REGION Network 2: Sterowanie grzałką w trybie automatycznym i manualnym
   // Gdy uruchomiony jest tryb automatyczny, wartość temperatury w szklarni powinna się mieścić w zakresie temperatury nastawionej +- wartość histerezy. Gdy jest ona za nieska uruchamiana jest grzałka. W trybie manualnym włączana jest ona od razu po naciśnięciu przycisku do niej przypisanego.
   RUNG wire#powerrail
      Contact( #czy_automatyczny )
      I_Contact( #czy_manualny )
      Sub(in1 := "Tryb_auto_parametry".Temperatura, in2 := #Wartosc_histerezy, out => #Histereza_minus)
      { S7_Templates := "SrcType := Real" } GT_Contact(in1 := #Histereza_minus, in2 := "Wejscia_PLC".Temperatura_wewnetrzna)
      wire#w1
      Coil( "Grzałka" )
   END_RUNG
   RUNG wire#powerrail
      Contact( #czy_manualny )
      I_Contact( #czy_automatyczny )
      Contact( "HMI".Przycisk_grzanie_manual )
   END_RUNG wire#w1
   // the same network as SCL:
   #_w1 := #czy_automatyczny AND NOT #czy_manualny;
   IF #_w1 THEN #Histereza_minus := "Tryb_auto_parametry".Temperatura - #Wartosc_histerezy; END_IF;
   "Grzałka" := (#_w1 AND (#Histereza_minus > "Wejscia_PLC".Temperatura_wewnetrzna)) OR (#czy_manualny AND NOT #czy_automatyczny AND "HMI".Przycisk_grzanie_manual);
END_REGION

REGION Network 3: TO DO Alarmy ostrzegające o nieosiąganiu wymaganej temperatury przez długi czas
   "IEC_Timer_0_DB_2".TON(IN := #czy_automatyczny AND NOT #czy_manualny AND ((#Histereza_plus < "Wejscia_PLC".Temperatura_wewnetrzna) OR (#Histereza_minus > "Wejscia_PLC".Temperatura_wewnetrzna)),
                          PT := T#30m);
   "Alarmy".Warning_wysoka_temp_1 := "IEC_Timer_0_DB_2".Q AND (#Histereza_plus > "Tryb_auto_parametry".Temperatura);
   "Alarmy".Warning_niska_temp_1 := "IEC_Timer_0_DB_2".Q AND (#Histereza_minus < "HMI".Temperatura_auto);
END_REGION
END_FUNCTION

FUNCTION "Zapis_parametrow_trybu_auto" : Void   // FC4, LAD
{ S7_Optimized_Access := 'TRUE' }
VERSION : 0.1
BEGIN

REGION Network 1: Zapis wybranych na HMI parametrów, aby zostały one stałe do kolejnego zatwierdzenia ich zmiany.
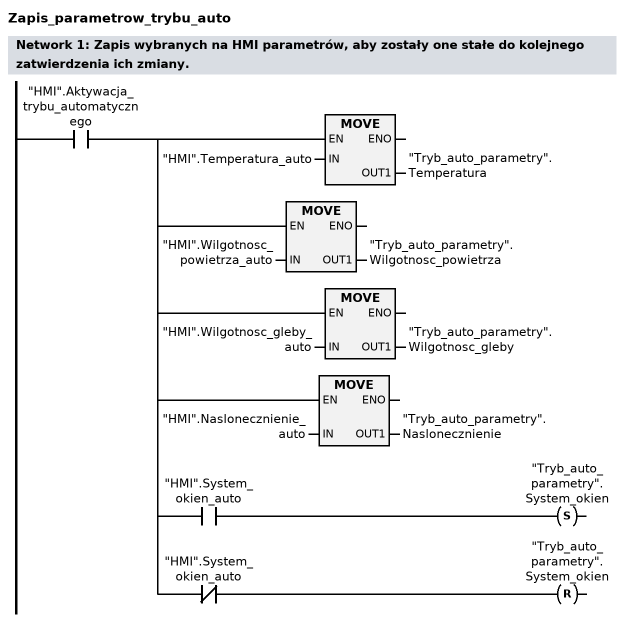
   RUNG wire#powerrail
      Contact( "HMI".Aktywacja_trybu_automatycznego )
      wire#w1
      Move(in := "HMI".Temperatura_auto, out1 => "Tryb_auto_parametry".Temperatura)
   END_RUNG
   RUNG wire#w1
      Move(in := "HMI".Wilgotnosc_powietrza_auto, out1 => "Tryb_auto_parametry".Wilgotnosc_powietrza)
   END_RUNG
   RUNG wire#w1
      Move(in := "HMI".Wilgotnosc_gleby_auto, out1 => "Tryb_auto_parametry".Wilgotnosc_gleby)
   END_RUNG
   RUNG wire#w1
      Move(in := "HMI".Naslonecznienie_auto, out1 => "Tryb_auto_parametry".Naslonecznienie)
   END_RUNG
   RUNG wire#w1
      Contact( "HMI".System_okien_auto )
      S_Coil( "Tryb_auto_parametry".System_okien )
   END_RUNG
   RUNG wire#w1
      I_Contact( "HMI".System_okien_auto )
      R_Coil( "Tryb_auto_parametry".System_okien )
   END_RUNG
   // the same network as SCL:
   IF "HMI".Aktywacja_trybu_automatycznego THEN
       "Tryb_auto_parametry".Temperatura := "HMI".Temperatura_auto;
       "Tryb_auto_parametry".Wilgotnosc_powietrza := "HMI".Wilgotnosc_powietrza_auto;
       "Tryb_auto_parametry".Wilgotnosc_gleby := "HMI".Wilgotnosc_gleby_auto;
       "Tryb_auto_parametry".Naslonecznienie := "HMI".Naslonecznienie_auto;
   END_IF;
   IF "HMI".Aktywacja_trybu_automatycznego AND "HMI".System_okien_auto THEN
       "Tryb_auto_parametry".System_okien := TRUE;
   END_IF;
   IF "HMI".Aktywacja_trybu_automatycznego AND NOT "HMI".System_okien_auto THEN
       "Tryb_auto_parametry".System_okien := FALSE;
   END_IF;
END_REGION
END_FUNCTION

FUNCTION "Jaki_Tryb" : Void   // FC5, LAD
{ S7_Optimized_Access := 'TRUE' }
VERSION : 0.1
BEGIN

REGION Network 1: Reset trybu auto jesli wykryje jakikolwiek inny tryb
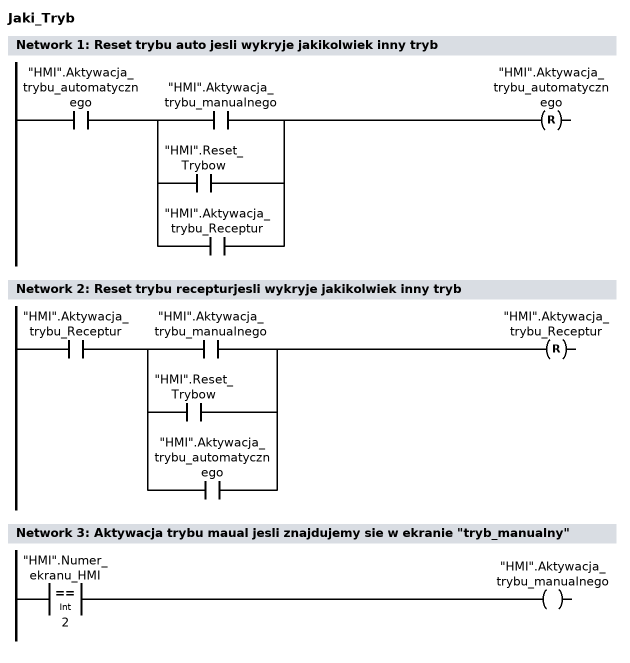
   RUNG wire#powerrail
      Contact( "HMI".Aktywacja_trybu_automatycznego )
      wire#w1
      Contact( "HMI".Aktywacja_trybu_manualnego )
      wire#w2
      R_Coil( "HMI".Aktywacja_trybu_automatycznego )
   END_RUNG
   RUNG wire#w1
      Contact( "HMI".Reset_Trybow )
   END_RUNG wire#w2
   RUNG wire#w1
      Contact( "HMI".Aktywacja_trybu_Receptur )
   END_RUNG wire#w2
   // the same network as SCL:
   IF "HMI".Aktywacja_trybu_automatycznego AND ("HMI".Aktywacja_trybu_manualnego OR "HMI".Reset_Trybow OR "HMI".Aktywacja_trybu_Receptur) THEN
       "HMI".Aktywacja_trybu_automatycznego := FALSE;
   END_IF;
END_REGION

REGION Network 2: Reset trybu recepturjesli wykryje jakikolwiek inny tryb
   RUNG wire#powerrail
      Contact( "HMI".Aktywacja_trybu_Receptur )
      wire#w1
      Contact( "HMI".Aktywacja_trybu_manualnego )
      wire#w2
      R_Coil( "HMI".Aktywacja_trybu_Receptur )
   END_RUNG
   RUNG wire#w1
      Contact( "HMI".Reset_Trybow )
   END_RUNG wire#w2
   RUNG wire#w1
      Contact( "HMI".Aktywacja_trybu_automatycznego )
   END_RUNG wire#w2
   // the same network as SCL:
   IF "HMI".Aktywacja_trybu_Receptur AND ("HMI".Aktywacja_trybu_manualnego OR "HMI".Reset_Trybow OR "HMI".Aktywacja_trybu_automatycznego) THEN
       "HMI".Aktywacja_trybu_Receptur := FALSE;
   END_IF;
END_REGION

REGION Network 3: Aktywacja trybu maual jesli znajdujemy sie w ekranie "tryb_manualny"
   RUNG wire#powerrail
      { S7_Templates := "SrcType := Int" } EQ_Contact(in1 := "HMI".Numer_ekranu_HMI, in2 := 2)
      Coil( "HMI".Aktywacja_trybu_manualnego )
   END_RUNG
   // the same network as SCL:
   "HMI".Aktywacja_trybu_manualnego := "HMI".Numer_ekranu_HMI = 2;
END_REGION
END_FUNCTION

FUNCTION "Ograniczanie_wartosci_parametrow" : Void   // FC6, LAD
TITLE = Każdy z poniższych network-ów odpowiada za to, aby po ustawieniu na HMI wartości przekraczajacej dopuszczalną, ta pozostała w wymaganym zakresie.
{ S7_Optimized_Access := 'TRUE' }
VERSION : 0.1
BEGIN

REGION Network 1: Ograniczenie dla wartosci ustawionej temperatury w trybie automatycznym
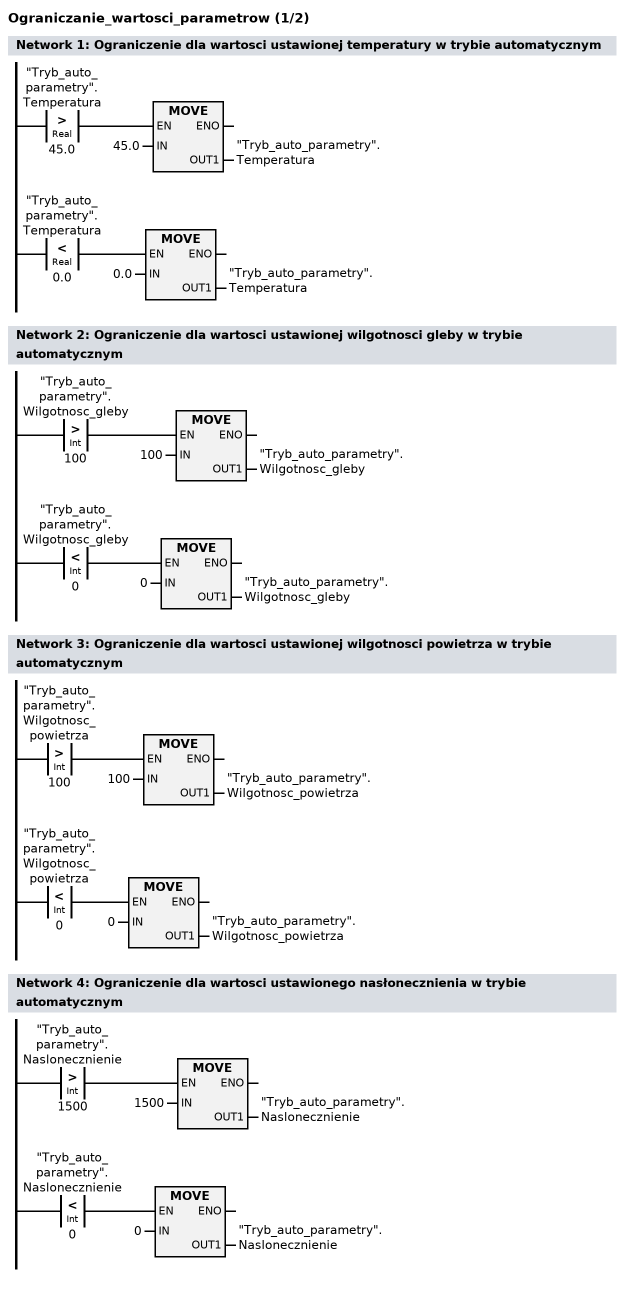
   RUNG wire#powerrail
      { S7_Templates := "SrcType := Real" } GT_Contact(in1 := "Tryb_auto_parametry".Temperatura, in2 := 45.0)
      Move(in := 45.0, out1 => "Tryb_auto_parametry".Temperatura)
   END_RUNG
   RUNG wire#powerrail
      { S7_Templates := "SrcType := Real" } LT_Contact(in1 := "Tryb_auto_parametry".Temperatura, in2 := 0.0)
      Move(in := 0.0, out1 => "Tryb_auto_parametry".Temperatura)
   END_RUNG
   // the same network as SCL:
   IF "Tryb_auto_parametry".Temperatura > 45.0 THEN "Tryb_auto_parametry".Temperatura := 45.0; END_IF;
   IF "Tryb_auto_parametry".Temperatura < 0.0 THEN "Tryb_auto_parametry".Temperatura := 0.0; END_IF;
END_REGION

REGION Network 2: Ograniczenie dla wartosci ustawionej wilgotnosci gleby w trybie automatycznym
   RUNG wire#powerrail
      { S7_Templates := "SrcType := Int" } GT_Contact(in1 := "Tryb_auto_parametry".Wilgotnosc_gleby, in2 := 100)
      Move(in := 100, out1 => "Tryb_auto_parametry".Wilgotnosc_gleby)
   END_RUNG
   RUNG wire#powerrail
      { S7_Templates := "SrcType := Int" } LT_Contact(in1 := "Tryb_auto_parametry".Wilgotnosc_gleby, in2 := 0)
      Move(in := 0, out1 => "Tryb_auto_parametry".Wilgotnosc_gleby)
   END_RUNG
   // the same network as SCL:
   IF "Tryb_auto_parametry".Wilgotnosc_gleby > 100 THEN
       "Tryb_auto_parametry".Wilgotnosc_gleby := 100;
   END_IF;
   IF "Tryb_auto_parametry".Wilgotnosc_gleby < 0 THEN "Tryb_auto_parametry".Wilgotnosc_gleby := 0; END_IF;
END_REGION

REGION Network 3: Ograniczenie dla wartosci ustawionej wilgotnosci powietrza w trybie automatycznym
   RUNG wire#powerrail
      { S7_Templates := "SrcType := Int" } GT_Contact(in1 := "Tryb_auto_parametry".Wilgotnosc_powietrza, in2 := 100)
      Move(in := 100, out1 => "Tryb_auto_parametry".Wilgotnosc_powietrza)
   END_RUNG
   RUNG wire#powerrail
      { S7_Templates := "SrcType := Int" } LT_Contact(in1 := "Tryb_auto_parametry".Wilgotnosc_powietrza, in2 := 0)
      Move(in := 0, out1 => "Tryb_auto_parametry".Wilgotnosc_powietrza)
   END_RUNG
   // the same network as SCL:
   IF "Tryb_auto_parametry".Wilgotnosc_powietrza > 100 THEN
       "Tryb_auto_parametry".Wilgotnosc_powietrza := 100;
   END_IF;
   IF "Tryb_auto_parametry".Wilgotnosc_powietrza < 0 THEN
       "Tryb_auto_parametry".Wilgotnosc_powietrza := 0;
   END_IF;
END_REGION

REGION Network 4: Ograniczenie dla wartosci ustawionego nasłonecznienia w trybie automatycznym
   RUNG wire#powerrail
      { S7_Templates := "SrcType := Int" } GT_Contact(in1 := "Tryb_auto_parametry".Naslonecznienie, in2 := 1500)
      Move(in := 1500, out1 => "Tryb_auto_parametry".Naslonecznienie)
   END_RUNG
   RUNG wire#powerrail
      { S7_Templates := "SrcType := Int" } LT_Contact(in1 := "Tryb_auto_parametry".Naslonecznienie, in2 := 0)
      Move(in := 0, out1 => "Tryb_auto_parametry".Naslonecznienie)
   END_RUNG
   // the same network as SCL:
   IF "Tryb_auto_parametry".Naslonecznienie > 1500 THEN
       "Tryb_auto_parametry".Naslonecznienie := 1500;
   END_IF;
   IF "Tryb_auto_parametry".Naslonecznienie < 0 THEN "Tryb_auto_parametry".Naslonecznienie := 0; END_IF;
END_REGION

REGION Network 5: Ograniczenie dla wartosci ustawionego stężenia CO2 w trybie automatycznym
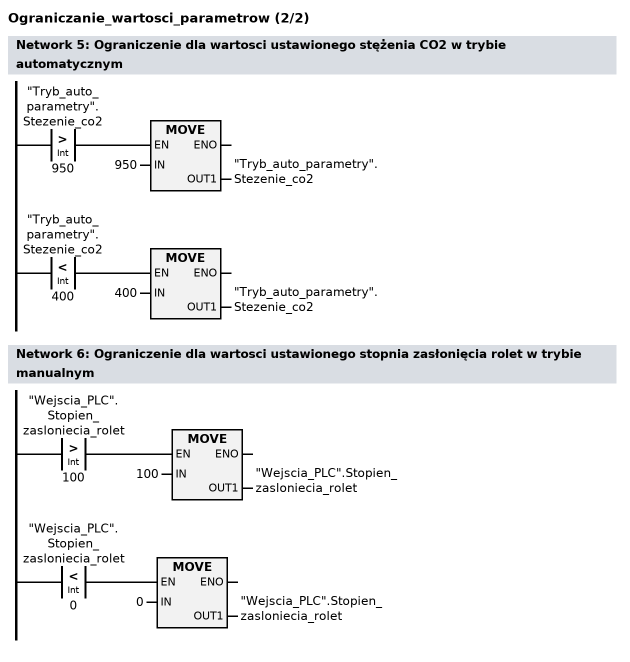
   RUNG wire#powerrail
      { S7_Templates := "SrcType := Int" } GT_Contact(in1 := "Tryb_auto_parametry".Stezenie_co2, in2 := 950)
      Move(in := 950, out1 => "Tryb_auto_parametry".Stezenie_co2)
   END_RUNG
   RUNG wire#powerrail
      { S7_Templates := "SrcType := Int" } LT_Contact(in1 := "Tryb_auto_parametry".Stezenie_co2, in2 := 400)
      Move(in := 400, out1 => "Tryb_auto_parametry".Stezenie_co2)
   END_RUNG
   // the same network as SCL:
   IF "Tryb_auto_parametry".Stezenie_co2 > 950 THEN "Tryb_auto_parametry".Stezenie_co2 := 950; END_IF;
   IF "Tryb_auto_parametry".Stezenie_co2 < 400 THEN "Tryb_auto_parametry".Stezenie_co2 := 400; END_IF;
END_REGION

REGION Network 6: Ograniczenie dla wartosci ustawionego stopnia zasłonięcia rolet w trybie manualnym
   RUNG wire#powerrail
      { S7_Templates := "SrcType := Int" } GT_Contact(in1 := "Wejscia_PLC".Stopien_zasloniecia_rolet, in2 := 100)
      Move(in := 100, out1 => "Wejscia_PLC".Stopien_zasloniecia_rolet)
   END_RUNG
   RUNG wire#powerrail
      { S7_Templates := "SrcType := Int" } LT_Contact(in1 := "Wejscia_PLC".Stopien_zasloniecia_rolet, in2 := 0)
      Move(in := 0, out1 => "Wejscia_PLC".Stopien_zasloniecia_rolet)
   END_RUNG
   // the same network as SCL:
   IF "Wejscia_PLC".Stopien_zasloniecia_rolet > 100 THEN
       "Wejscia_PLC".Stopien_zasloniecia_rolet := 100;
   END_IF;
   IF "Wejscia_PLC".Stopien_zasloniecia_rolet < 0 THEN "Wejscia_PLC".Stopien_zasloniecia_rolet := 0; END_IF;
END_REGION
END_FUNCTION

FUNCTION "Sterowanie_podlewaniem_zraszaniem" : Void   // FC7, LAD
{ S7_Optimized_Access := 'TRUE' }
VERSION : 0.1
   VAR_INPUT
      Czy_automatyczny : Bool;
      Czy_manualny : Bool;
   END_VAR
BEGIN

REGION Network 1: Sterowanie pompą zraszaczy, które odpowiadają za wilgotność powietrza w szklarni
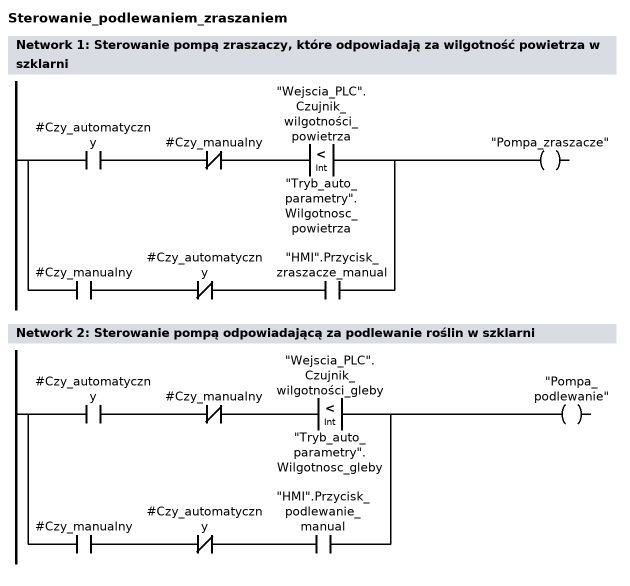
   RUNG wire#powerrail
      Contact( #Czy_automatyczny )
      I_Contact( #Czy_manualny )
      { S7_Templates := "SrcType := Int" } LT_Contact(in1 := "Wejscia_PLC".Czujnik_wilgotności_powietrza, in2 := "Tryb_auto_parametry".Wilgotnosc_powietrza)
      wire#w1
      Coil( "Pompa_zraszacze" )
   END_RUNG
   RUNG wire#powerrail
      Contact( #Czy_manualny )
      I_Contact( #Czy_automatyczny )
      Contact( "HMI".Przycisk_zraszacze_manual )
   END_RUNG wire#w1
   // the same network as SCL:
   "Pompa_zraszacze" := (#Czy_automatyczny AND NOT #Czy_manualny AND ("Wejscia_PLC".Czujnik_wilgotności_powietrza < "Tryb_auto_parametry".Wilgotnosc_powietrza)) OR (#Czy_manualny AND NOT #Czy_automatyczny AND "HMI".Przycisk_zraszacze_manual);
END_REGION

REGION Network 2: Sterowanie pompą odpowiadającą za podlewanie roślin w szklarni
   RUNG wire#powerrail
      Contact( #Czy_automatyczny )
      I_Contact( #Czy_manualny )
      { S7_Templates := "SrcType := Int" } LT_Contact(in1 := "Wejscia_PLC".Czujnik_wilgotności_gleby, in2 := "Tryb_auto_parametry".Wilgotnosc_gleby)
      wire#w1
      Coil( "Pompa_podlewanie" )
   END_RUNG
   RUNG wire#powerrail
      Contact( #Czy_manualny )
      I_Contact( #Czy_automatyczny )
      Contact( "HMI".Przycisk_podlewanie_manual )
   END_RUNG wire#w1
   // the same network as SCL:
   "Pompa_podlewanie" := (#Czy_automatyczny AND NOT #Czy_manualny AND ("Wejscia_PLC".Czujnik_wilgotności_gleby < "Tryb_auto_parametry".Wilgotnosc_gleby)) OR (#Czy_manualny AND NOT #Czy_automatyczny AND "HMI".Przycisk_podlewanie_manual);
END_REGION
END_FUNCTION

FUNCTION "Sterowanie_oknami" : Void   // FC8, LAD
{ S7_Optimized_Access := 'TRUE' }
VERSION : 0.1
   VAR_INPUT
      czy_manualny : Bool;
      czy_automatyczny : Bool;
   END_VAR
   VAR_TEMP
      Histereza_plus : Int;
      Histereza_minus : Int;
      Zakres_temp_gora : Real;   // Górny zakres temperatury zewnętrznej dla której w trybie automatycznym będą otwierane okna
      Zakres_temp_dol : Real;   // Dolny zakres temperatury zewnętrznej dla której w trybie automatycznym będą otwierane okna
   END_VAR
   VAR CONSTANT
      Histereza : Int := 25;   // Histereza, która określa kiedy stan CO2 w szklarni jest uznawany za prawidłowy
   END_VAR
BEGIN

REGION Network 1: Operacje matematyczne używane w networku 2. i 3.
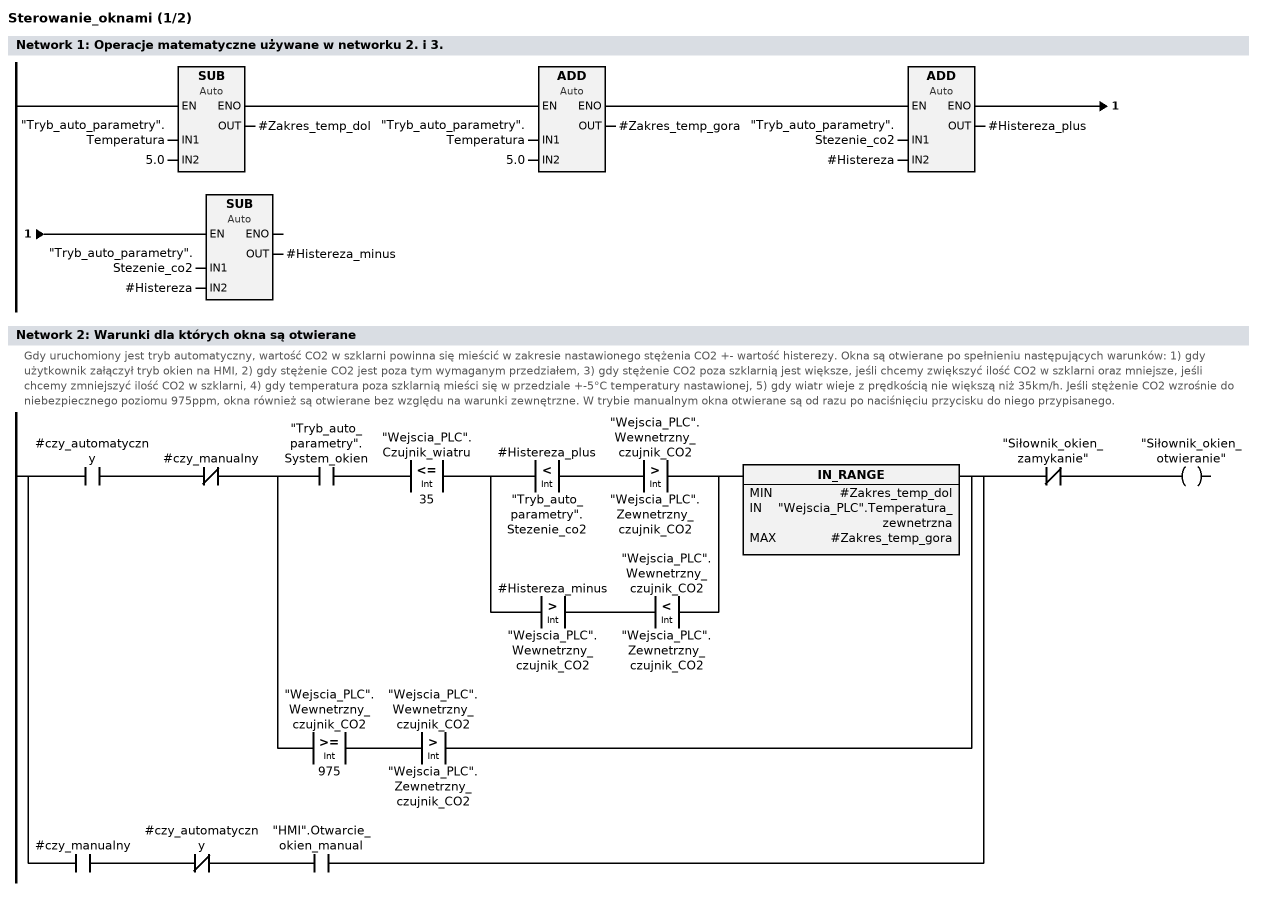
   RUNG wire#powerrail
      Sub(in1 := "Tryb_auto_parametry".Temperatura, in2 := 5.0, out => #Zakres_temp_dol)
      Add(in1 := "Tryb_auto_parametry".Temperatura, in2 := 5.0, out => #Zakres_temp_gora)
      Add(in1 := "Tryb_auto_parametry".Stezenie_co2, in2 := #Histereza, out => #Histereza_plus)
      Sub(in1 := "Tryb_auto_parametry".Stezenie_co2, in2 := #Histereza, out => #Histereza_minus)
   END_RUNG
   // the same network as SCL:
   #Zakres_temp_dol := "Tryb_auto_parametry".Temperatura - 5.0;
   #Zakres_temp_gora := "Tryb_auto_parametry".Temperatura + 5.0;
   #Histereza_plus := "Tryb_auto_parametry".Stezenie_co2 + #Histereza;
   #Histereza_minus := "Tryb_auto_parametry".Stezenie_co2 - #Histereza;
END_REGION

REGION Network 2: Warunki dla których okna są otwierane
   // Gdy uruchomiony jest tryb automatyczny, wartość CO2 w szklarni powinna się mieścić w zakresie nastawionego stężenia CO2 +- wartość histerezy. Okna są otwierane po spełnieniu następujących warunków: 1) gdy użytkownik załączył tryb okien na HMI, 2) gdy stężenie CO2 jest poza tym wymaganym przedziałem, 3) gdy stężenie CO2 poza szklarnią jest większe, jeśli chcemy zwiększyć ilość CO2 w szklarni oraz mniejsze, jeśli chcemy zmniejszyć ilość CO2 w szklarni, 4) gdy temperatura poza szklarnią mieści się w przedziale +-5°C temperatury nastawionej, 5) gdy wiatr wieje z prędkością nie większą niż 35km/h. Jeśli stężenie CO2 wzrośnie do niebezpiecznego poziomu 975ppm, okna również są otwierane bez względu na warunki zewnętrzne. W trybie manualnym okna otwierane są od razu po naciśnięciu przycisku do niego przypisanego.
   RUNG wire#powerrail
      Contact( #czy_automatyczny )
      I_Contact( #czy_manualny )
      wire#w1
      Contact( "Tryb_auto_parametry".System_okien )
      { S7_Templates := "SrcType := Int" } LE_Contact(in1 := "Wejscia_PLC".Czujnik_wiatru, in2 := 35)
      wire#w2
      { S7_Templates := "SrcType := Int" } LT_Contact(in1 := #Histereza_plus, in2 := "Tryb_auto_parametry".Stezenie_co2)
      { S7_Templates := "SrcType := Int" } GT_Contact(in1 := "Wejscia_PLC".Wewnetrzny_czujnik_CO2, in2 := "Wejscia_PLC".Zewnetrzny_czujnik_CO2)
      wire#w3
      { S7_Templates := "SrcType := Real" } InRange(min := #Zakres_temp_dol, in := "Wejscia_PLC".Temperatura_zewnetrzna, max := #Zakres_temp_gora)
      wire#w4
      I_Contact( "Siłownik_okien_zamykanie" )
      Coil( "Siłownik_okien_otwieranie" )
   END_RUNG
   RUNG wire#w2
      { S7_Templates := "SrcType := Int" } GT_Contact(in1 := #Histereza_minus, in2 := "Wejscia_PLC".Wewnetrzny_czujnik_CO2)
      { S7_Templates := "SrcType := Int" } LT_Contact(in1 := "Wejscia_PLC".Wewnetrzny_czujnik_CO2, in2 := "Wejscia_PLC".Zewnetrzny_czujnik_CO2)
   END_RUNG wire#w3
   RUNG wire#w1
      { S7_Templates := "SrcType := Int" } GE_Contact(in1 := "Wejscia_PLC".Wewnetrzny_czujnik_CO2, in2 := 975)
      { S7_Templates := "SrcType := Int" } GT_Contact(in1 := "Wejscia_PLC".Wewnetrzny_czujnik_CO2, in2 := "Wejscia_PLC".Zewnetrzny_czujnik_CO2)
   END_RUNG wire#w4
   RUNG wire#powerrail
      Contact( #czy_manualny )
      I_Contact( #czy_automatyczny )
      Contact( "HMI".Otwarcie_okien_manual )
   END_RUNG wire#w4
   // the same network as SCL:
   "Siłownik_okien_otwieranie" := ((#czy_automatyczny AND NOT #czy_manualny AND (("Tryb_auto_parametry".System_okien AND ("Wejscia_PLC".Czujnik_wiatru <= 35) AND (((#Histereza_plus < "Tryb_auto_parametry".Stezenie_co2) AND ("Wejscia_PLC".Wewnetrzny_czujnik_CO2 > "Wejscia_PLC".Zewnetrzny_czujnik_CO2)) OR ((#Histereza_minus > "Wejscia_PLC".Wewnetrzny_czujnik_CO2) AND ("Wejscia_PLC".Wewnetrzny_czujnik_CO2 < "Wejscia_PLC".Zewnetrzny_czujnik_CO2))) AND (#Zakres_temp_dol <= "Wejscia_PLC".Temperatura_zewnetrzna) AND ("Wejscia_PLC".Temperatura_zewnetrzna <= #Zakres_temp_gora)) OR (("Wejscia_PLC".Wewnetrzny_czujnik_CO2 >= 975) AND ("Wejscia_PLC".Wewnetrzny_czujnik_CO2 > "Wejscia_PLC".Zewnetrzny_czujnik_CO2)))) OR (#czy_manualny AND NOT #czy_automatyczny AND "HMI".Otwarcie_okien_manual)) AND NOT "Siłownik_okien_zamykanie";
END_REGION

REGION Network 3: Warunki dla których okna są zamykane
   // W trybie automatycznym okna są zamykane: 1) gdy tryb okien został wyłączony przez użytkownika, 2) gdy stężenie CO2 w szklarni wynosi zadaną wartość tego parametru +- histereza, 3) gdy stężenie CO2 poza szklarnią jest mniejsze, niż wewnątrz, jeśli chcemy zwiększyć jego ilość oraz większe, gdy chcemy zmniejszyć jego ilość, 4) gdy tempperatura zewnętrzna różni się o ponad 5°C od zadanej, 5) gdy wiatr wieje z prędkością większą niż 35km/h, 6) gdy stężenie CO2 w szklarni nie przekracza 955ppm lub przekracza, ale stężenie CO2 poza szklarnią jest większe. W trybie manualnym okna są zamykane, gdy przełączk na HMI znajdzie się w pozycji "ZAMKNIĘTE".
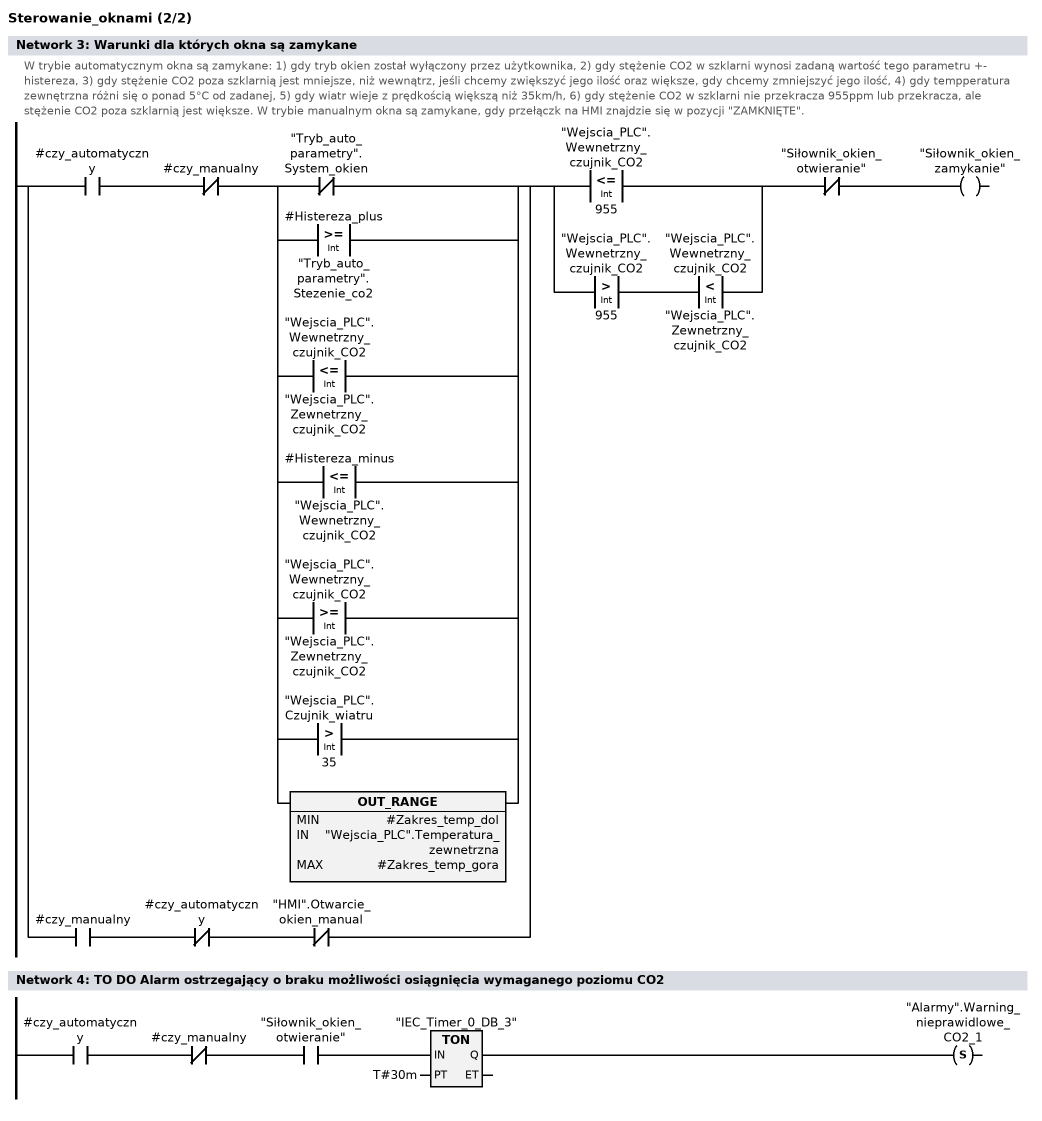
   "Siłownik_okien_zamykanie" := ((#czy_automatyczny AND NOT #czy_manualny AND (NOT "Tryb_auto_parametry".System_okien OR (#Histereza_plus >= "Tryb_auto_parametry".Stezenie_co2) OR ("Wejscia_PLC".Wewnetrzny_czujnik_CO2 <= "Wejscia_PLC".Zewnetrzny_czujnik_CO2) OR (#Histereza_minus <= "Wejscia_PLC".Wewnetrzny_czujnik_CO2) OR ("Wejscia_PLC".Wewnetrzny_czujnik_CO2 >= "Wejscia_PLC".Zewnetrzny_czujnik_CO2) OR ("Wejscia_PLC".Czujnik_wiatru > 35) OR ("Wejscia_PLC".Temperatura_zewnetrzna < #Zakres_temp_dol) OR ("Wejscia_PLC".Temperatura_zewnetrzna > #Zakres_temp_gora))) OR (#czy_manualny AND NOT #czy_automatyczny AND NOT "HMI".Otwarcie_okien_manual)) AND (("Wejscia_PLC".Wewnetrzny_czujnik_CO2 <= 955) OR (("Wejscia_PLC".Wewnetrzny_czujnik_CO2 > 955) AND ("Wejscia_PLC".Wewnetrzny_czujnik_CO2 < "Wejscia_PLC".Zewnetrzny_czujnik_CO2))) AND NOT "Siłownik_okien_otwieranie";
END_REGION

REGION Network 4: TO DO Alarm ostrzegający o braku możliwości osiągnięcia wymaganego poziomu CO2
   "IEC_Timer_0_DB_3".TON(IN := #czy_automatyczny AND NOT #czy_manualny AND "Siłownik_okien_otwieranie",
                          PT := T#30m);
   IF "IEC_Timer_0_DB_3".Q THEN "Alarmy".Warning_nieprawidlowe_CO2_1 := TRUE; END_IF;
END_REGION
END_FUNCTION

FUNCTION "SYMULACJA" : Void   // FC9, LAD
{ S7_Optimized_Access := 'TRUE' }
VERSION : 0.1
   VAR_INPUT
      counters : Bool;
   END_VAR
   VAR_TEMP
      temperatura_temp : Real;
      roznica_temperatur : Real;
      "wilgotność powietrza_temp" : Int;
      wilgotnosc_gleby_temp : Int;
      stezenie_CO2 : Int;
      natezenie_swiatla_temp : Int;
      odsloniecie_okna_temp : Real;
      pedkosc_wiatru_temp : Real;
      rand : Real;
      error : Bool;
      status : Int;
      sub_status : Int;
      rolety_temp : Real;
      test1 : Real;
   END_VAR
   VAR_TEMP   // added for the SCL form of the ladder/FBD networks
      _w1 : Bool;
   END_VAR
BEGIN

REGION Network 1: blok oblicza roznice temperatur
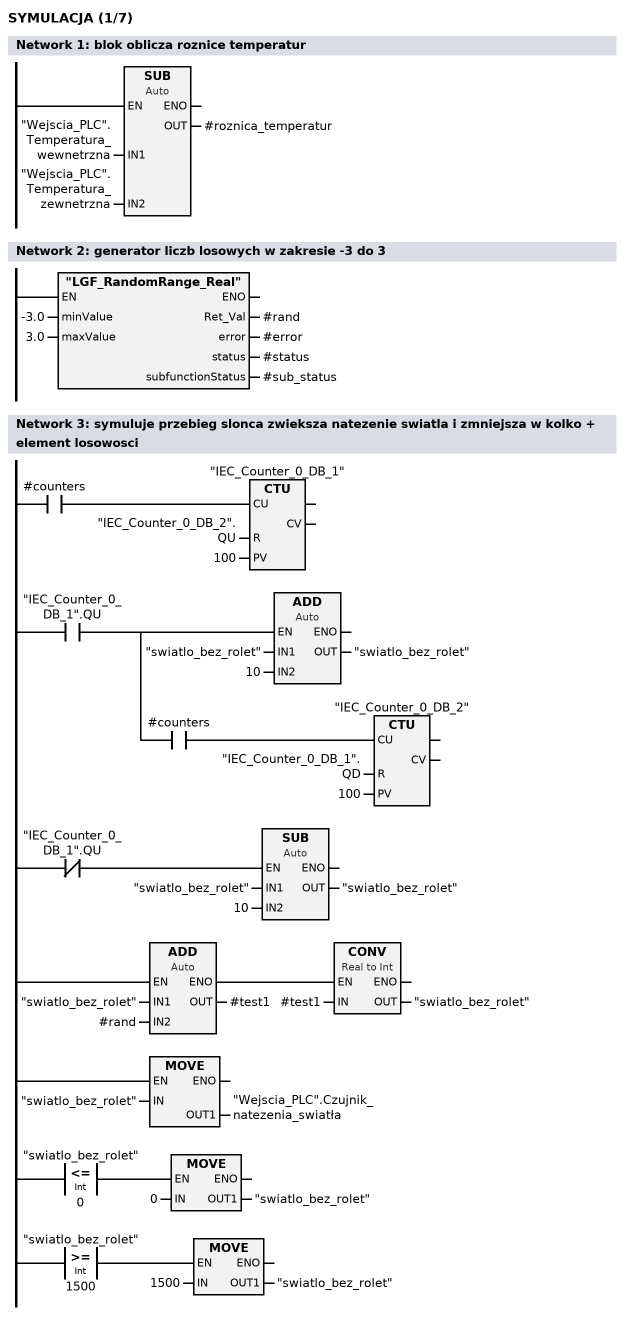
   RUNG wire#powerrail
      { S7_GenerateENO := "TRUE" } Sub(in1 := "Wejscia_PLC".Temperatura_wewnetrzna, in2 := "Wejscia_PLC".Temperatura_zewnetrzna, out => #roznica_temperatur)
   END_RUNG
   // the same network as SCL:
   #roznica_temperatur := "Wejscia_PLC".Temperatura_wewnetrzna - "Wejscia_PLC".Temperatura_zewnetrzna;
END_REGION

REGION Network 2: generator liczb losowych w zakresie -3 do 3
   RUNG wire#powerrail
      "LGF_RandomRange_Real"(minValue := -3.0, maxValue := 3.0, Ret_Val => #rand, error => #error, status => #status, subfunctionStatus => #sub_status)
   END_RUNG
   // the same network as SCL:
   #rand := "LGF_RandomRange_Real"(minValue := -3.0,
                           maxValue := 3.0,
                           error => #error,
                           status => #status,
                           subfunctionStatus => #sub_status);
END_REGION

REGION Network 3: symuluje przebieg slonca zwieksza natezenie swiatla i zmniejsza w kolko + element losowosci
   // ENO of a box is taken as its EN; it also drops when the box reports an error
   "IEC_Counter_0_DB_1".CTU(CU := #counters, R := "IEC_Counter_0_DB_2".QU, PV := 100);
   IF "IEC_Counter_0_DB_1".QU THEN "swiatlo_bez_rolet" := "swiatlo_bez_rolet" + 10; END_IF;
   "IEC_Counter_0_DB_2".CTU(CU := "IEC_Counter_0_DB_1".QU AND #counters,
                           R := "IEC_Counter_0_DB_1".QD,
                           PV := 100);
   IF NOT "IEC_Counter_0_DB_1".QU THEN "swiatlo_bez_rolet" := "swiatlo_bez_rolet" - 10; END_IF;
   #test1 := "swiatlo_bez_rolet" + #rand;
   "swiatlo_bez_rolet" := REAL_TO_INT(#test1);
   "Wejscia_PLC".Czujnik_natezenia_swiatła := "swiatlo_bez_rolet";
   IF "swiatlo_bez_rolet" <= 0 THEN "swiatlo_bez_rolet" := 0; END_IF;
   IF "swiatlo_bez_rolet" >= 1500 THEN "swiatlo_bez_rolet" := 1500; END_IF;
END_REGION

REGION Network 4: funkcja oblicza liniową zależność natężenia światła od zasłonięcia rolet
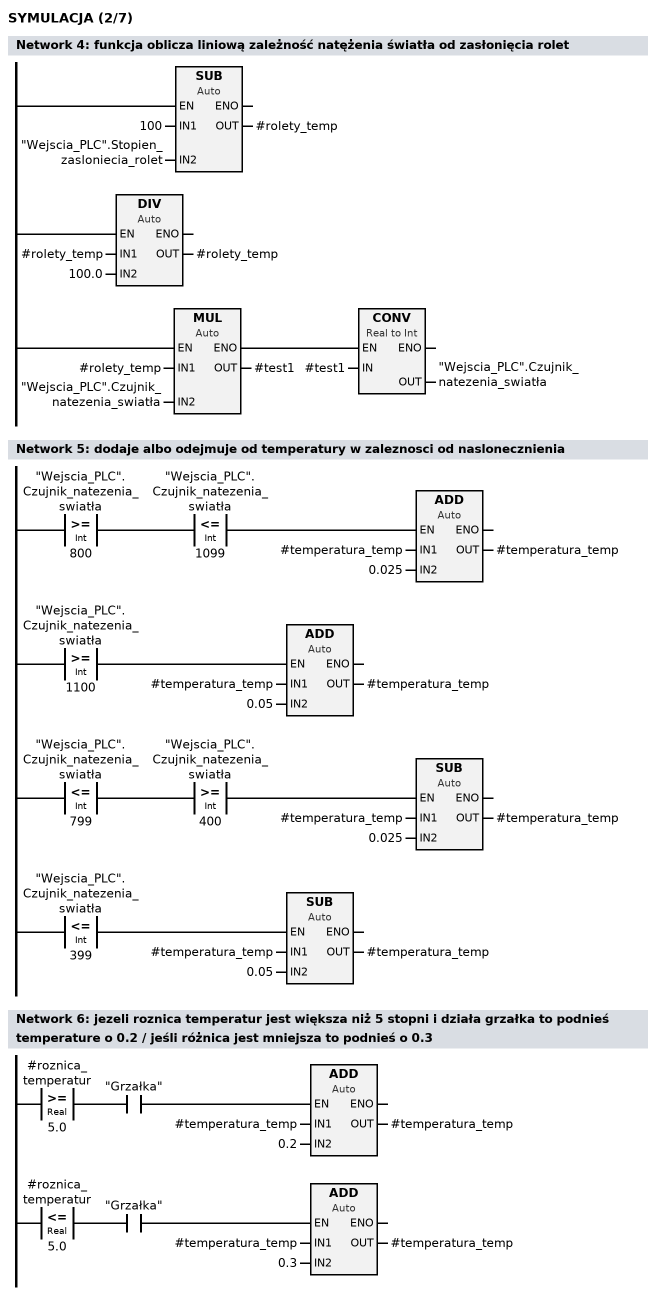
   RUNG wire#powerrail
      { S7_GenerateENO := "TRUE" } Sub(in1 := 100, in2 := "Wejscia_PLC".Stopien_zasloniecia_rolet, out => #rolety_temp)
   END_RUNG
   RUNG wire#powerrail
      { S7_GenerateENO := "TRUE" } Div(in1 := #rolety_temp, in2 := 100.0, out => #rolety_temp)
   END_RUNG
   RUNG wire#powerrail
      { S7_GenerateENO := "TRUE" } Mul(in1 := #rolety_temp, in2 := "Wejscia_PLC".Czujnik_natezenia_swiatła, out => #test1)
      { S7_Templates := "[SrcType := Real, DestType := Int]"; S7_GenerateENO := "TRUE" } Convert(in := #test1, out => "Wejscia_PLC".Czujnik_natezenia_swiatła)
   END_RUNG
   // the same network as SCL:
   // ENO of a box is taken as its EN; it also drops when the box reports an error
   #rolety_temp := 100 - "Wejscia_PLC".Stopien_zasloniecia_rolet;
   #rolety_temp := #rolety_temp / 100.0;
   #test1 := #rolety_temp * "Wejscia_PLC".Czujnik_natezenia_swiatła;
   "Wejscia_PLC".Czujnik_natezenia_swiatła := REAL_TO_INT(#test1);
END_REGION

REGION Network 5: dodaje albo odejmuje od temperatury w zaleznosci od naslonecznienia
   RUNG wire#powerrail
      { S7_Templates := "SrcType := Int" } GE_Contact(in1 := "Wejscia_PLC".Czujnik_natezenia_swiatła, in2 := 800)
      { S7_Templates := "SrcType := Int" } LE_Contact(in1 := "Wejscia_PLC".Czujnik_natezenia_swiatła, in2 := 1099)
      { S7_GenerateENO := "TRUE" } Add(in1 := #temperatura_temp, in2 := 0.025, out => #temperatura_temp)
   END_RUNG
   RUNG wire#powerrail
      { S7_Templates := "SrcType := Int" } GE_Contact(in1 := "Wejscia_PLC".Czujnik_natezenia_swiatła, in2 := 1100)
      { S7_GenerateENO := "TRUE" } Add(in1 := #temperatura_temp, in2 := 0.05, out => #temperatura_temp)
   END_RUNG
   RUNG wire#powerrail
      { S7_Templates := "SrcType := Int" } LE_Contact(in1 := "Wejscia_PLC".Czujnik_natezenia_swiatła, in2 := 799)
      { S7_Templates := "SrcType := Int" } GE_Contact(in1 := "Wejscia_PLC".Czujnik_natezenia_swiatła, in2 := 400)
      { S7_GenerateENO := "TRUE" } Sub(in1 := #temperatura_temp, in2 := 0.025, out => #temperatura_temp)
   END_RUNG
   RUNG wire#powerrail
      { S7_Templates := "SrcType := Int" } LE_Contact(in1 := "Wejscia_PLC".Czujnik_natezenia_swiatła, in2 := 399)
      { S7_GenerateENO := "TRUE" } Sub(in1 := #temperatura_temp, in2 := 0.05, out => #temperatura_temp)
   END_RUNG
   // the same network as SCL:
   IF ("Wejscia_PLC".Czujnik_natezenia_swiatła >= 800) AND ("Wejscia_PLC".Czujnik_natezenia_swiatła <= 1099) THEN
       #temperatura_temp := #temperatura_temp + 0.025;
   END_IF;
   IF "Wejscia_PLC".Czujnik_natezenia_swiatła >= 1100 THEN
       #temperatura_temp := #temperatura_temp + 0.05;
   END_IF;
   IF ("Wejscia_PLC".Czujnik_natezenia_swiatła <= 799) AND ("Wejscia_PLC".Czujnik_natezenia_swiatła >= 400) THEN
       #temperatura_temp := #temperatura_temp - 0.025;
   END_IF;
   IF "Wejscia_PLC".Czujnik_natezenia_swiatła <= 399 THEN
       #temperatura_temp := #temperatura_temp - 0.05;
   END_IF;
END_REGION

REGION Network 6: jezeli roznica temperatur jest większa niż 5 stopni i działa grzałka to podnieś temperature o 0.2 / jeśli różnica jest mniejsza to podnieś o 0.3
   RUNG wire#powerrail
      { S7_Templates := "SrcType := Real" } GE_Contact(in1 := #roznica_temperatur, in2 := 5.0)
      Contact( "Grzałka" )
      { S7_GenerateENO := "TRUE" } Add(in1 := #temperatura_temp, in2 := 0.2, out => #temperatura_temp)
   END_RUNG
   RUNG wire#powerrail
      { S7_Templates := "SrcType := Real" } LE_Contact(in1 := #roznica_temperatur, in2 := 5.0)
      Contact( "Grzałka" )
      { S7_GenerateENO := "TRUE" } Add(in1 := #temperatura_temp, in2 := 0.3, out => #temperatura_temp)
   END_RUNG
   // the same network as SCL:
   IF (#roznica_temperatur >= 5.0) AND "Grzałka" THEN #temperatura_temp := #temperatura_temp + 0.2; END_IF;
   IF (#roznica_temperatur <= 5.0) AND "Grzałka" THEN #temperatura_temp := #temperatura_temp + 0.3; END_IF;
END_REGION

REGION Network 7: jezeli działa wentylator to obniż temperature o 0.1
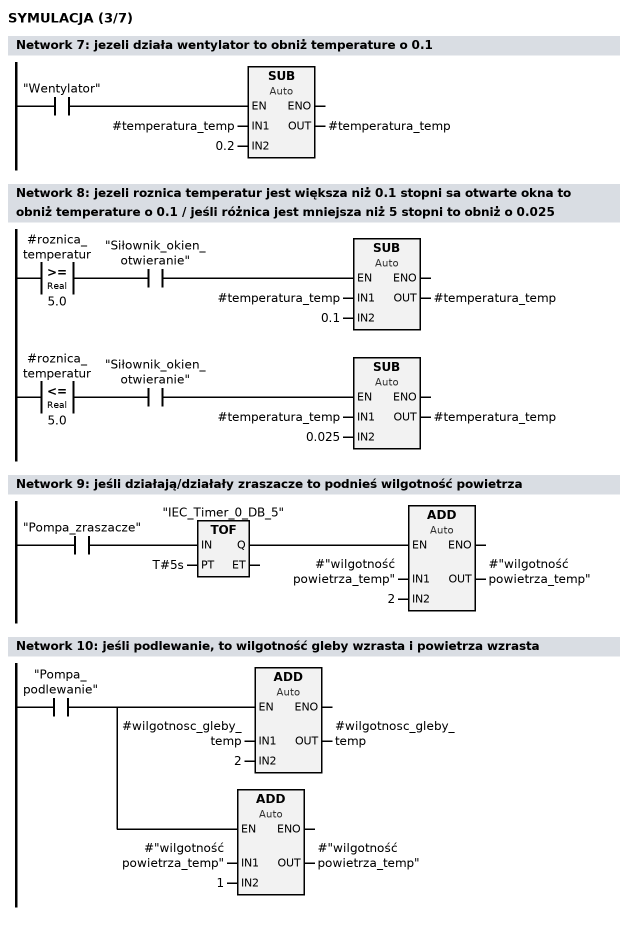
   RUNG wire#powerrail
      Contact( "Wentylator" )
      { S7_GenerateENO := "TRUE" } Sub(in1 := #temperatura_temp, in2 := 0.2, out => #temperatura_temp)
   END_RUNG
   // the same network as SCL:
   IF "Wentylator" THEN #temperatura_temp := #temperatura_temp - 0.2; END_IF;
END_REGION

REGION Network 8: jezeli roznica temperatur jest większa niż 0.1 stopni sa otwarte okna to obniż temperature o 0.1 / jeśli różnica jest mniejsza niż 5 stopni to obniż o 0.025
   RUNG wire#powerrail
      { S7_Templates := "SrcType := Real" } GE_Contact(in1 := #roznica_temperatur, in2 := 5.0)
      Contact( "Siłownik_okien_otwieranie" )
      { S7_GenerateENO := "TRUE" } Sub(in1 := #temperatura_temp, in2 := 0.1, out => #temperatura_temp)
   END_RUNG
   RUNG wire#powerrail
      { S7_Templates := "SrcType := Real" } LE_Contact(in1 := #roznica_temperatur, in2 := 5.0)
      Contact( "Siłownik_okien_otwieranie" )
      { S7_GenerateENO := "TRUE" } Sub(in1 := #temperatura_temp, in2 := 0.025, out => #temperatura_temp)
   END_RUNG
   // the same network as SCL:
   IF (#roznica_temperatur >= 5.0) AND "Siłownik_okien_otwieranie" THEN
       #temperatura_temp := #temperatura_temp - 0.1;
   END_IF;
   IF (#roznica_temperatur <= 5.0) AND "Siłownik_okien_otwieranie" THEN
       #temperatura_temp := #temperatura_temp - 0.025;
   END_IF;
END_REGION

REGION Network 9: jeśli działają/działały zraszacze to podnieś wilgotność powietrza
   "IEC_Timer_0_DB_5".TOF(IN := "Pompa_zraszacze", PT := T#5s);
   IF "IEC_Timer_0_DB_5".Q THEN #"wilgotność powietrza_temp" := #"wilgotność powietrza_temp" + 2; END_IF;
END_REGION

REGION Network 10: jeśli podlewanie, to wilgotność gleby wzrasta i powietrza wzrasta
   RUNG wire#powerrail
      Contact( "Pompa_podlewanie" )
      wire#w1
      { S7_GenerateENO := "TRUE" } Add(in1 := #wilgotnosc_gleby_temp, in2 := 2, out => #wilgotnosc_gleby_temp)
   END_RUNG
   RUNG wire#w1
      { S7_GenerateENO := "TRUE" } Add(in1 := #"wilgotność powietrza_temp", in2 := 1, out => #"wilgotność powietrza_temp")
   END_RUNG
   // the same network as SCL:
   IF "Pompa_podlewanie" THEN
       #wilgotnosc_gleby_temp := #wilgotnosc_gleby_temp + 2;
       #"wilgotność powietrza_temp" := #"wilgotność powietrza_temp" + 1;
   END_IF;
END_REGION

REGION Network 11: realizacja zaleznosci odslaniania i zaslaniania rolet, od stopnia zasłonięcia